(* Logix 5000 project; controller PLC_MCC1300_75F1 vendor 1 type 14 code 166 rev 32.11; software revision 32.04; part 60 of 83 *)
(* tags used below, declared in another part *)
   CM_ConveyorStackerToLine_JS1_Sync : CM_ConveyorStackerToLine;
   CONST_dDest_Cullet : DINT;
   CONST_dDest_Stk : DINT;
   CONST_rgdDestMask : DINT[32];   // Destination Mask
   Convoy_SL_DATA_NULL : UDT_Convoy_SL;
   GP_CheckIdPlatePresent : GP_CheckIdPlatePresent;
   GP_InvertCapxLite : GP_InvertCapxLite;
   GP_OB_InitializeMain : GP_OB_Initialize;
   GP_RampSpace : GP_RampSpace;
   Gp_SpaceConvUtilities_V1 : GP_SpaceConvUtilities_V1;
   M310Popup : MAC_Popup_ZC[2];
   M311 : MAC_Conveyor;
   M311_Data : UDT_Convoy_SL;
   M311_SpaceConv_Utilities : SpaceConv_Utilities;
   M312 : MAC_Conveyor_Single;
   M315A_SpaceConv_Utilities : SpaceConv_Utilities;
   M315A_SpaceConvUtilities : SpaceConv_Utilities;
   M315B : MAC_Conveyor;
   M315B_ALM : MAC_Conveyor_ALM;
   M315B_Data : UDT_Convoy_SL;
   M315B_HMW : MAC_Conveyor_HMW;
   M315B_SpaceConv_Utilities : SpaceConv_Utilities;
   M315B_xPlateCullet : BOOL;
   M315Popup : MAC_Popup_ZC[2];
   M315Popup_SL_DATA : UDT_Convoy_SL;
   TMP_d : DINT;
   TMP_dConveyorNumberForZoneCleaning : DINT;
   TMP_dDecelerationPositionEndConveyor : DINT;
   TMP_dHeadPosition : DINT;
   TMP_dOffsetLoadUnload_cmm : DINT;
   TMP_dPhEndPosition_cmm : DINT;
   TMP_dTailPosition : DINT;
   TMP_rgxId : DINT[10];
   TMP_SendToCullet : BOOL;
   TMP_xConveyorInvolvedInCleaning : BOOL;
   TMP_xConveyorOfStartCleaning : BOOL;
   TMP_xCulletPresent : BOOL;
   TMP_xEnableLoadUnload : BOOL;
   TMP_xEnableZoneCleaning : BOOL;
   TMP_xLiteThisDestPresent : BOOL;
   TMP_xReqUnpack : BOOL;
   xAlwaysOFF : BOOL;
   xAlwaysON : BOOL;
   xDebugOFF : BOOL;
   Z402 : MAC_Zone;
   Z402_HMR : MAC_Zone_HMR;
   Z402_HMW : MAC_Zone_HMW;
(* MainProgram, continued *)

ROUTINE M315B_Alarm   (* ladder *)
   // Reset Alarm
   0: XIC(Z402.tmON_ResetAlarm.DN)FLL(0,M315B_ALM,1);
   1: XIC(Z402.ST_xEnableControlError)XIC(M315B.INPUT_xDriveError_M2)OTL(M315B_ALM.rgxStoppingFault_M[0].11);
   2: XIC(Z402.ST_xEnableControlError)XIO(M315B.INPUT_xDriveError_M2)[XIC(M315B.OUTPUT_xRun_M2) ,XIC(M315B.OUTPUT_xReverse_M2) ,XIC(M315B.OUTPUT_xPositioning_M2) ]XIO(M315B.INPUT_xDriveFeedback_M2)[XIO(M315B.tmON_FeedbackTimeOut_M2.DN) TON(M315B.tmON_FeedbackTimeOut_M2,?,?) ,XIC(M315B.tmON_FeedbackTimeOut_M2.DN) OTL(M315B_ALM.rgxStoppingFault_M[0].12) ];
   3: XIC(Z402.ST_xEnableControlError)XIO(M315B.INPUT_xMotorThermalProbe_M2)XIC(xDebugOFF)OTL(M315B_ALM.rgxStoppingFault_M[0].14);
   4: XIC(Z402.ST_xEnableControlError)[XIC(M315B.INPUT_xDriveInhibit_M2) ,XIC(M315B.OUTPUT_xDriveEnable_M2) XIO(M315B.INPUT_xDriveReady_M2) ][XIO(M315B.tmON_DriveInhibit_M2.DN) TON(M315B.tmON_DriveInhibit_M2,?,?) ,XIC(M315B.tmON_DriveInhibit_M2.DN) OTL(M315B_ALM.rgxStoppingFault_M[0].16) ];
   5: XIC(Z402.ST_xEnableControlError)XIC(M315B.INPUT_xDriveError_M1)OTL(M315B_ALM.rgxStoppingFault_M[0].1);
   6: XIC(Z402.ST_xEnableControlError)XIO(M315B.INPUT_xDriveError_M1)[XIC(M315B.OUTPUT_xRun_M1) ,XIC(M315B.OUTPUT_xReverse_M1) ,XIC(M315B.OUTPUT_xPositioning_M1) ]XIO(M315B.INPUT_xDriveFeedback_M1)[XIO(M315B.tmON_FeedbackTimeOut_M1.DN) TON(M315B.tmON_FeedbackTimeOut_M1,?,?) ,XIC(M315B.tmON_FeedbackTimeOut_M1.DN) OTL(M315B_ALM.rgxStoppingFault_M[0].2) ];
   7: XIC(Z402.ST_xEnableControlError)XIO(M315B.INPUT_xMotorThermalProbe_M1)XIC(xDebugOFF)OTL(M315B_ALM.rgxStoppingFault_M[0].4);
   8: XIC(Z402.ST_xEnableControlError)[XIC(M315B.INPUT_xDriveInhibit_M1) ,XIC(M315B.OUTPUT_xDriveEnable_M1) XIO(M315B.INPUT_xDriveReady_M1) ][XIO(M315B.tmON_DriveInhibit_M1.DN) TON(M315B.tmON_DriveInhibit_M1,?,?) ,XIC(M315B.tmON_DriveInhibit_M1.DN) OTL(M315B_ALM.rgxStoppingFault_M[0].6) ];
   9: XIC(M315B.ST_xEnableControlError)XIC(M315B.PH_x.7)NEQ(M315B_SpaceConv_Utilities.CONST_dSyncMode,0)[XIO(M315B.ST_xPlateSynchronized) OTL(M315B_ALM.rgxWarning[0].0) ,XIC(M315B.ST_xPlateSynchronized) OTU(M315B_ALM.rgxWarning[0].0) ];
   10: XIC(M315B.ST_xEnableControlError)XIC(M315B.PH_x.7)[XIC(M315B_Data.tFlag.tConveyor.xReqStop) ,XIC(M315B_Data.tFlag.tConveyor.xBypassReqEndStop) ]OTL(M315B_ALM.rgxWarning[0].1);
   // #####_CUMULATIVE ALARM_#####
   11: NOP();
   12: [NEQ(M315B_ALM.rgxStoppingFault[0],0) ,NEQ(M315B_ALM.rgxStoppingFault_M[0],0) ,NEQ(M315B_ALM.rgxStoppingFault_M[1],0) ]OTE(M315B.ST_xStopMachineFault);
   13: [NEQ(M315B_ALM.rgxFault[0],0) ,NEQ(M315B_ALM.rgxFault_M[0],0) ,NEQ(M315B_ALM.rgxFault_M[1],0) ]OTE(M315B.ST_xStopNextCycleFault);
END_ROUTINE

ROUTINE M315B_Logic   (* ladder *)
   // #####_COSTANTS_#####
   0: [MOV(3100,TMP_dConveyorNumberForZoneCleaning) MOV(50000,TMP_dOffsetLoadUnload_cmm) MOV(500,M315B_SpaceConv_Utilities.CONST_dPresetFeedbackTime_ms) OTU(TMP_xEnableLoadUnload) OTU(TMP_xEnableZoneCleaning) MOV(485000,M315B_SpaceConv_Utilities.CONST_dConveyorLength_cmm) MOV(375000,M315B_SpaceConv_Utilities.CONST_dConveyorWidth_cmm) SUB(M315B_SpaceConv_Utilities.CONST_dConveyorLength_cmm,30000,M315B.AUX_dPresetStopLoad_cmm) ADD(M315B_SpaceConv_Utilities.CONST_dConveyorLength_cmm,90000,M315B.AUX_dPresetStopUnload_cmm) MOV(1.2,M315B_SpaceConv_Utilities.CONST_rAcceleration_ms2) MOV(1.2,M315B_SpaceConv_Utilities.CONST_rDeceleration_ms2) MOV(M315B_SpaceConv_Utilities.CONST_dConveyorLength_cmm,TMP_dPhEndPosition_cmm) ,XIC(M315B.PH_x.28) [MOV(1,M315B_SpaceConv_Utilities.CONST_dSyncMode) ,MUL(M315B_SpaceConv_Utilities.CONST_dSyncroPhPosition_cmm,-1,M315B_SpaceConv_Utilities.CONST_dSyncroPhPosition_cmm) ,MOV(200000,M315B_SpaceConv_Utilities.CONST_dSyncroPhWindow_cmm) ] ];
   // #####_MATCH_#####
   1: NOP();
   // Conveyor Cleaning
   2: XIC(TMP_xEnableZoneCleaning)XIC(Z402.ST_xCleaningAccepted)GRT(Z402_HMW.dCleaningSelection,0)[EQU(Z402_HMW.dCleaningSelection,TMP_dConveyorNumberForZoneCleaning) OTE(TMP_xConveyorOfStartCleaning) ,GEQ(Z402_HMW.dCleaningSelection,TMP_dConveyorNumberForZoneCleaning) OTE(TMP_xConveyorInvolvedInCleaning) ];
   // Enable control error
   3: XIC(Z402.ST_xEnableControlError)OTE(M315B.ST_xEnableControlError);
   // Mode 7 - Offsett for load/unload Simultaney
   4: XIC(M315B.PH_x.8)MOV(M315B.AUX_dPresetStopLoad_cmm,M315B_SpaceConv_Utilities.ST_dStopLoadForseen_cmm)MOV(TMP_dOffsetLoadUnload_cmm,M315B_SpaceConv_Utilities.CONF_MD7_dOffset_cmm)GP_SpaceConvUtilities_V1(Gp_SpaceConvUtilities_V1,M315B_SpaceConv_Utilities,M315B_SpaceConv_Utilities,M315A_SpaceConvUtilities,7);
   // #####_ALARMS_#####
   5: NOP();
   // Call Alarm Routine
   6: JSR(M315B_Alarm,0);
   // #####_HMI_LOGICS_#####
   7: NOP();
   // Condition ok for Cleaning
   8: [XIO(TMP_xEnableZoneCleaning) ,XIC(TMP_xEnableZoneCleaning) XIC(M315B.ST_xOutputEnable) [XIO(TMP_xConveyorOfStartCleaning) ,XIC(M315B.PH_x.0) ,XIO(M315B.PH_x.8) ] ]OTE(M315B.ST_xCleaningConditionOK);
   // Cleaning Accepted
   9: [[XIC(M315B_HMW.xStopLocalCleaningRequest) ,XIC(Z402_HMW.xStopCleanZoneRequest) ] OTU(M315B_HMW.xStopLocalCleaningRequest) OTU(M315B_HMW.xLocalCleaningRequest) ,[XIC(M315B_HMW.xLocalCleaningRequest) ,XIC(Z402.ST_xCleaningAccepted) ] [XIC(M315B.ST_xCleaningConditionOK) ,XIC(M315B.ST_xCleaningAccepted) ] OTE(M315B.ST_xCleaningAccepted) ];
   // Manual Mode Enabled
   10: XIO(M315B_SpaceConv_Utilities.ST_xFeedbackRotation)[XIC(M315B_HMW.xEnableDisableManualCommand) XIC(M315B.ST_xConditionOKStopCycle) OTL(M315B.ST_xManualMode) ,XIO(M315B_HMW.xEnableDisableManualCommand) OTU(M315B.ST_xManualMode) ];
   // Virtual door enabled
   11: XIC(M315B_HMW.xEnableDisableVirtualDoor)OTE(M315B.ST_xVirtualDoorEnabled);
   // Clear manual command
   12: XIO(M315B.ST_xManualMode)MOV(0,M315B_HMW.rgxMan);
   // #####_STATUSES_#####
   13: NOP();
   // Syncro  -  OS Syncro Photocell
   14: XIC(xAlwaysON)[XIC(M315B.INPUT_xSyncroPhotocell_1) ONS(M315B.OSR_xSynchroPhotocellHead) OTE(M315B.OS_xSynchroPhotocellHead) GEQ(M315B_SpaceConv_Utilities.CONST_dSyncMode,1) OTE(M315B_SpaceConv_Utilities.ST_OS_xSynchroPhotocellHead) ,XIO(M315B.INPUT_xSyncroPhotocell_1) ONS(M315B.OSR_xSynchroPhotocellTail) OTE(M315B.OS_xSynchroPhotocellTail) GEQ(M315B_SpaceConv_Utilities.CONST_dSyncMode,2) OTE(M315B_SpaceConv_Utilities.ST_OS_xSynchroPhotocellTail) ];
   // Id Plate presence
   15: MOV(CONST_rgdDestMask[24],CONST_dDest_Cullet)GP_CheckIdPlatePresent(GP_CheckIdPlatePresent,M315B_Data,TMP_rgxId,M315B.ST_xIdPlatePresence,TMP_xCulletPresent,CONST_dDest_Cullet)MOV(CONST_rgdDestMask[0],CONST_dDest_Stk)GP_CheckIdPlatePresent(GP_CheckIdPlatePresent,M315B_Data,TMP_rgxId,M315B.ST_xIdPlatePresence,TMP_xLiteThisDestPresent,CONST_dDest_Stk)XIC(TMP_xCulletPresent)OTE(M315B_xPlateCullet);
   // Machine in Alarm
   16: [XIC(M315B.ST_xStopMachineFault) ,XIC(M315B.ST_xStopNextCycleFault) ]OTE(M315B.ST_xMachineAlarm);
   // Condition ok for stop Cycle
   17: [XIO(M315B.ST_xPhasesInProgress) ,XIC(M315B.PH_x.8) XIO(M315B.OUTPUT_xRun_M1) XIO(M315B.OUTPUT_xRun_M2) XIO(M315B_SpaceConv_Utilities.ST_xFeedbackRotation) ,XIC(M315B.PH_x.9) XIO(M315B.OUTPUT_xRun_M1) XIO(M315B_SpaceConv_Utilities.ST_xFeedbackRotation) ,XIC(M315B.ST_xMachineAlarm) ,XIO(Z402.ST_xCycleON) ]OTE(M315B.ST_xConditionOKStopCycle);
   // Cycle load unload simultaneous
   18: XIC(TMP_xEnableLoadUnload)XIO(M315B.ST_xDisableLoadUnloadOnStop)XIO(M315B.ST_xIdPlatePresence)OTE(M315B.ST_xCycleLoadUnload);
   // Speed Management
   19: [XIO(M315B_SpaceConv_Utilities.O_xRampInProgress) XIO(M315B.ST_xManualMode) MOV(Z402_HMR.dLineSpeed_mm_min,M315B.AUX_dReqSpeed_mm_min) ,XIC(M315B.ST_xManualMode) MOV(Z402_HMW.dManualSpeed_mm_min,M315B.AUX_dReqSpeed_mm_min) ,NEQ(M315B.AUX_dReqSpeed_mm_min,M315B_SpaceConv_Utilities.ST_dRealSpeed_mm_min) OTE(M315B.OS_xChangeSpeed) ];
   // Ramp Management
   20: GP_RampSpace(GP_RampSpace,M315B_SpaceConv_Utilities.CONST_rAcceleration_ms2,M315B_SpaceConv_Utilities.CONST_rDeceleration_ms2,M315B_SpaceConv_Utilities.ST_dRealSpeed_mm_min,M315B.AUX_dAccSpace_cmm,M315B.AUX_dDecSpace_cmm);
   // Space Convoy utilities MOD 1 for Calculate Head/Tail
   21: XIC(xAlwaysON)[[XIC(M315B.OUTPUT_xRun_M1) ,XIC(M315B.OUTPUT_xReverse_M1) ] XIO(M315B.ST_xManualMode) OTE(M315B_SpaceConv_Utilities.CONF_MD1_xRun) ,XIC(M315B.OUTPUT_xReverse_M1) XIC(xAlwaysOFF) XIO(M315B.ST_xManualMode) OTE(M315B_SpaceConv_Utilities.CONF_MD1_xReverse) ,[XIC(M315B.INPUT_xDriveFeedback_M1) ,XIC(M315B_SpaceConv_Utilities.CONF_MD1_xRun) GRT(M315B_SpaceConv_Utilities.O_dCountFeedbackTime_ms,0) ] OTE(M315B_SpaceConv_Utilities.ST_xFeedbackRotation) ,XIC(M315B.ST_xIdPlatePresence) OTE(M315B_SpaceConv_Utilities.CONF_MD1_xHeadTracking) ,XIC(M315B.ST_xPlatePresence) OTE(M315B_SpaceConv_Utilities.CONF_MD1_xTailTracking) ,MOV(GP_OB_InitializeMain.OUT_dExecutionTime_ms,M315B_SpaceConv_Utilities.CONF_MD1_dScan_ms) GP_SpaceConvUtilities_V1(Gp_SpaceConvUtilities_V1,M315B_SpaceConv_Utilities,M315B_SpaceConv_Utilities,M315A_SpaceConv_Utilities,1) ];
   // Output Enable
   22: XIC(Z402.ST_xCycleON)XIO(M315B.ST_xManualMode)XIO(M315B.ST_xStopMachineFault)[XIO(M315B.ST_xPlatePassageUpstream_FW) XIO(M315B.ST_xPlatePassageUpstream_BKW) ,XIC(M315B.ST_xPlatePassageUpstream_BKW) XIC(M311.ST_xOutputEnable) ][XIC(M315B.INPUT_xHighPositionPopup_1) ,XIC(M315B.INPUT_xHighPositionPopup_2) ]OTE(M315B.ST_xOutputEnable);
   23: GRT(M315B_Data.dTotalCaps,1)OTE(TMP_xReqUnpack);
   // #####_WORKING_FLAGS_#####
   24: NOP();
   // #####_LOGICS_#####
   25: NOP();
   // Phase of load
   26: XIC(xAlwaysOFF)[OTL(M315B.PH_x.0) ,OTU(M315B_SpaceConv_Utilities.O_xPlateSynchronized) ,OTU(M315B.ST_xDisableLoadUnloadOnStop) ,OTE(M315B.OS_xLoad_FW) ,COP(M315B_Data,M315B_Data,1) FLL(0,M315B_Data,1) ,GP_SpaceConvUtilities_V1(Gp_SpaceConvUtilities_V1,M315B_SpaceConv_Utilities,M315B_SpaceConv_Utilities,M315A_SpaceConv_Utilities,5) ];
   // Syncro  -  Space Convoy utilities MOD 4
   27: GRT(M315B_SpaceConv_Utilities.CONST_dSyncMode,0)[[XIC(M315B.PH_x.0) XIO(M315B.PH_x.8) ,XIC(M315B.PH_x.1) XIO(M315B.PH_x.9) ] ,[XIC(M315B.PH_x.0) XIC(M315B.PH_x.8) ,XIC(M315B.PH_x.1) XIC(M315B.PH_x.9) ] ADD(M315B_SpaceConv_Utilities.CONST_dSyncroPhPosition_cmm,TMP_dOffsetLoadUnload_cmm,TMP_d) GRT(M315B_SpaceConv_Utilities.O_dTailPosition_cmm,TMP_d) ][MOV(M315B_Data.dLength_cmm,M315B_SpaceConv_Utilities.CONF_MD4_MD6_dLength_cmm) ,GP_SpaceConvUtilities_V1(Gp_SpaceConvUtilities_V1,M315B_SpaceConv_Utilities,M315B_SpaceConv_Utilities,M315A_SpaceConv_Utilities,4) ];
   // End load Phase
   28: XIC(M315B.PH_x.0)GRT(M315B_SpaceConv_Utilities.O_dHeadPosition_cmm,M315B.AUX_dPresetStopLoad_cmm)[OTE(M315B.PH_x.7) ,OTU(M315B.PH_x.0) ,OTL(M315B.ST_xPlatePresence) ];
   // End load Phase
   29: XIC(M315B.PH_x.1)GRT(M315B_SpaceConv_Utilities.O_dHeadPosition_cmm,M315B.AUX_dPresetStopLoad_cmm)[OTE(M315B.PH_x.5) ,OTU(M315B.PH_x.1) ,OTL(M315B.ST_xPlatePresence) ];
   // New data received from MainLine
   30: XIC(M315B.ST_xAux4)XIC(M310Popup[0].ST_xPlateDataReadyToSend)XIC(M310Popup[0].PH_xEndRise)[GP_InvertCapxLite(GP_InvertCapxLite,0,1,1,M315Popup_SL_DATA,M315B_Data,Convoy_SL_DATA_NULL,M315B_SpaceConv_Utilities.CONST_dConveyorWidth_cmm,M315B_SpaceConv_Utilities.CONST_dConveyorLength_cmm,M315B_SpaceConv_Utilities.CONF_MD2_MD3_dPrstPos_cmm,M315Popup[0].AUX_dReqTarget_cmm,200000) ,GP_SpaceConvUtilities_V1(Gp_SpaceConvUtilities_V1,M315B_SpaceConv_Utilities,M315B_SpaceConv_Utilities,M315B_SpaceConv_Utilities,2) ,OTL(M315B.ST_xPlatePresence) ];
   31: XIC(M315B.ST_xAux4)XIC(M310Popup[0].ST_xPlateDataReadyToSend)XIC(M310Popup[0].PH_xEndRise)GRT(M315B_Data.dTotalCaps,1)MOV(30000,M315B_Data.rgtCap[0].dReqGapForConv_cmm)MOV(30000,M315B_Data.rgtCap[1].dReqGapForConv_cmm)[XIC(xAlwaysOFF) SUB(M315B_SpaceConv_Utilities.O_dHeadPosition_cmm,50000,TMP_dHeadPosition) ,XIO(xAlwaysOFF) SUB(M315B_Data.dLength_cmm,20000,TMP_dHeadPosition) ]SUB(TMP_dHeadPosition,M315B_Data.dLength_cmm,TMP_dTailPosition);
   // Calculation Space for Wait Stop Next Conveyor
   32: CPT(TMP_dDecelerationPositionEndConveyor,M315B_SpaceConv_Utilities.CONST_dConveyorLength_cmm - M315B.AUX_dAccSpace_cmm + 1000);
   // Wait stop next Machine
   33: XIO(M315B.PH_x.8)XIO(M315B.PH_x.9)XIO(M315B.PH_x.10)GEQ(M315B_SpaceConv_Utilities.O_dHeadPosition_cmm,TMP_dDecelerationPositionEndConveyor)OTE(M315B.ST_xWaitStopNextMachine);
   // Set Wait Machine Stop
   34: [[XIC(M315B.PH_x.7) ,XIC(M315B.PH_x.5) ] [XIO(M311.ST_xInitialConditionOK) ,XIC(M315B.ST_xWaitStopNextMachine) [XIC(M311_SpaceConv_Utilities.O_xRampInProgress) ,XIO(M311_SpaceConv_Utilities.ST_xFeedbackRotation) ] ] ,[XIC(M315B.PH_x.0) ,XIC(M315B.PH_x.1) ] NEQ(Z402_HMR.dLineSpeed_mm_min,M315B.AUX_dReqSpeed_mm_min) ]OTL(M315B.ST_xWaitMachineStop);
   // Reset Wait Machine Stop
   35: XIO(M315B_SpaceConv_Utilities.ST_xFeedbackRotation)[XIO(M315B_SpaceConv_Utilities.ST_xFeedbackRotation) ,XIO(M315B.ST_xWaitStopNextMachine) ]EQU(Z402_HMR.dLineSpeed_mm_min,M315B.AUX_dReqSpeed_mm_min)OTU(M315B.ST_xWaitMachineStop);
   // Unpack management
   // -
   // -
   36: NOP();
   // Phase of unpacking
   37: XIC(Z402.ST_xConditionOkPhaseAdvancement)XIC(M315B.ST_xPlatePresence)XIC(M315B.ST_xIdPlatePresence)XIC(M315B.ST_xOutputEnable)XIC(M311.ST_xInitialConditionOK)XIO(M315B.ST_xWaitMachineStop)XIO(M315B.ST_xPhasesInProgress)XIC(TMP_xReqUnpack)XIC(TMP_xLiteThisDestPresent)[XIC(M315B.ST_xAxleReadyToMoveDelayed) ,XIC(xAlwaysON) ][OTL(M315B.PH_x.16) ,XIO(M315B.PH_x.16) OTL(M315B.PH_x.18) ,[XIC(M315B.PH_x.16) ,XIC(M315B.PH_x.18) ] OTE(M315B.OS_xUnpack) ,MOV(M315B_Data.dLength_cmm,M315B_SpaceConv_Utilities.CONF_MD4_MD6_dLength_cmm) GP_SpaceConvUtilities_V1(Gp_SpaceConvUtilities_V1,M315B_SpaceConv_Utilities,M315B_SpaceConv_Utilities,M315A_SpaceConv_Utilities,6) ,MOV(M315B_Data.rgtCap[0].dLength_cmm,M315B.AUX_dPhPosTarget_cmm) ];
   38: XIC(Z402.ST_xConditionOkPhaseAdvancement)XIC(M315B.ST_xOutputEnable)XIC(M315B.ST_xPlatePresence)XIC(M315B.ST_xIdPlatePresence)XIO(M315B.ST_xWaitMachineStop)XIO(M315B.ST_xPhasesInProgress)OTE(M315B.ST_xWaitReadyToMove);
   // Phase of unload
   39: XIC(Z402.ST_xConditionOkPhaseAdvancement)XIC(TMP_xLiteThisDestPresent)XIC(M315B.ST_xPlatePresence)XIC(M315B.ST_xIdPlatePresence)XIO(TMP_xReqUnpack)XIC(M315B.ST_xOutputEnable)XIC(M311.ST_xInitialConditionOK)XIO(M315B.ST_xWaitMachineStop)XIO(M315B.ST_xPhasesInProgress)[XIC(M315B.ST_xAxleReadyToMoveDelayed) ,XIC(xAlwaysON) ]XIC(TMP_xLiteThisDestPresent)XIO(M315B.PH_x.8)[OTL(M315B.PH_x.8) ,OTE(M315B.OS_xUnload_FW) ,MOV(M315B_Data.dLength_cmm,M315B_SpaceConv_Utilities.CONF_MD4_MD6_dLength_cmm) GP_SpaceConvUtilities_V1(Gp_SpaceConvUtilities_V1,M315B_SpaceConv_Utilities,M315B_SpaceConv_Utilities,M315A_SpaceConv_Utilities,6) ];
   // Phase of end unload
   40: XIC(M315B.PH_x.8)[[GEQ(M315B_SpaceConv_Utilities.O_dTailPosition_cmm,M315B.AUX_dPresetStopUnload_cmm) ,XIC(M311.PH_x.7) ] ,XIO(M315B_SpaceConv_Utilities.ST_xFeedbackRotation) GEQ(M315B_SpaceConv_Utilities.O_dTailPosition_cmm,M315B_SpaceConv_Utilities.CONST_dConveyorLength_cmm) ][OTE(M315B.PH_x.15) ,OTU(M315B.PH_x.8) ,OTU(M315B.ST_xPlatePresence) ];
   // Stop for unload on main line
   41: XIC(Z402.ST_xConditionOkPhaseAdvancement)XIC(M315B.INPUT_xHighPositionPopup_1)XIC(M315B.INPUT_xHighPositionPopup_2)XIC(M315B.ST_xOutputEnable)XIO(M315B.ST_xPhasesInProgress)XIC(M315B.ST_xPlatePresence)XIC(M315B.ST_xIdPlatePresence)XIO(TMP_xLiteThisDestPresent)[OTL(M315B.PH_x.22) ,GP_InvertCapxLite(GP_InvertCapxLite,1,0,1,M315B_Data,M315Popup_SL_DATA,Convoy_SL_DATA_NULL,M315B_SpaceConv_Utilities.CONST_dConveyorLength_cmm,M315B_SpaceConv_Utilities.CONST_dConveyorWidth_cmm,M315B_SpaceConv_Utilities.CONF_MD2_MD3_dPrstPos_cmm,M315B_SpaceConv_Utilities.O_dHeadPosition_cmm,225000) ];
   // End stop for unload on main line
   42: XIC(M315B.PH_x.22)XIO(M315B.INPUT_xHighPositionPopup_1)XIO(M315B.INPUT_xHighPositionPopup_2)[OTU(M315B.PH_x.22) ,OTE(M315B.PH_x.23) ,OTU(M315B.ST_xPlatePresence) ,FLL(0,M315B_Data,1) ];
   // Phase in progress
   43: NEQ(M315B.PH_x,0)OTE(M315B.ST_xPhasesInProgress);
   // #####_CLEANING_#####
   44: NOP();
   // Cleaning Reset
   45: [XIC(M315B.ST_xCleaningAccepted) [XIC(Z402.ST_xCleaningAccepted) ,XIO(TMP_xConveyorOfStartCleaning) ] ,XIC(M315B.INPUT_xLowPositionPopup_1) XIC(M315B.INPUT_xLowPositionPopup_2) ][XIC(M315B.ST_xIdPlatePresence) OTL(TMP_SendToCullet) FLL(0,M315B_Data,1) ,MOV(0,M315B.PH_x) OTU(M315B.ST_xPlatePresence) ];
   // Initial condition OK (to main line)
   46: XIC(Z402.ST_xConditionOkPhaseAdvancement)XIC(Z402.ST_xCycleON)XIO(M315B.ST_xManualMode)XIO(M315B.ST_xStopMachineFault)XIO(M315B_HMW.xEnableDisableManualCommand)XIO(M315B.ST_xReqCleaning)XIO(M315B.ST_xCleaningAccepted)XIO(M315B_HMW.xLocalCleaningRequest)XIO(M315B.ST_xStopNextCycleFault)XIO(M315B.ST_xVirtualDoorEnabled)XIO(M315B.ST_xPhasesInProgress)XIO(M315B.ST_xPlatePresence)XIO(M311.ST_xAux1)XIO(M312.ST_xAux1)XIO(CM_ConveyorStackerToLine_JS1_Sync.xRequestReturnInLine)XIO(CM_ConveyorStackerToLine_JS1_Sync.xRotationForUnload)OTE(M315B.ST_xAux4);
   // #### Plate reentry ####
   47: NOP();
   // Initial condition reentry
   48: XIC(Z402.ST_xConditionOkPhaseAdvancement)XIC(M315B.ST_xOutputEnable)XIC(M315B.INPUT_xHighPositionPopup_1)XIC(M315B.INPUT_xHighPositionPopup_2)XIO(M315B_HMW.xEnableDisableManualCommand)XIO(M315B.ST_xReqCleaning)XIO(M315B.ST_xCleaningAccepted)XIO(M315B.ST_xStopNextCycleFault)XIO(M311.ST_xVirtualDoorEnabled)XIO(M315B.ST_xPhasesInProgress)XIO(M315B.ST_xPlatePresence)XIO(M315B.ST_xIdPlatePresence)OTE(M315B.ST_xInitialConditionOK_BW);
   // Phase of load
   49: XIC(M311.OS_xUnload_BW)[XIC(M311.PH_x.24) OTL(M315B.PH_x.28) ,COP(M311_Data,M315B_Data,1) FLL(0,M311_Data,1) ,OTU(M315B_SpaceConv_Utilities.ST_xLastModLoadBkw) ,GP_SpaceConvUtilities_V1(Gp_SpaceConvUtilities_V1,M315B_SpaceConv_Utilities,M315B_SpaceConv_Utilities,M315A_SpaceConv_Utilities,15) ];
